REGION Network 357
   RUNG wire#powerrail
      Contact( "DuplicateCarrierfound" )
      Coil( "Carrier_17_Duplicate_Carrier_Fault" )
   END_RUNG
   // the same network as SCL:
   "Carrier_17_Duplicate_Carrier_Fault" := "DuplicateCarrierfound";
END_REGION

REGION Network 358
   RUNG wire#powerrail
      Contact( "EMS".Carrier[17].SDC_OUT.Faults.MotionOnFault )
      Coil( "Carrier_17_Motion_On_Fault" )
   END_RUNG
   // the same network as SCL:
   "Carrier_17_Motion_On_Fault" := "EMS".Carrier[17].SDC_OUT.Faults.MotionOnFault;
END_REGION

REGION Network 359
   RUNG wire#powerrail
      Contact( "EMS".Carrier[17].SDC_OUT.Faults.MotionOffFault )
      Coil( "Carrier_17_Motion_Off_Fault" )
   END_RUNG
   // the same network as SCL:
   "Carrier_17_Motion_Off_Fault" := "EMS".Carrier[17].SDC_OUT.Faults.MotionOffFault;
END_REGION

REGION Network 360
   RUNG wire#powerrail
      Contact( "EMS".Carrier[17].SDC_OUT.Faults.CarrierSpacingFault )
      Coil( "Carrier_17_Carrier_Spacing_Fault" )
   END_RUNG
   // the same network as SCL:
   "Carrier_17_Carrier_Spacing_Fault" := "EMS".Carrier[17].SDC_OUT.Faults.CarrierSpacingFault;
END_REGION

REGION Network 361
   RUNG wire#powerrail
      Move(in := "EMS".Carrier[18].SDC_OUT.Zone, out1 => "Carrier_18_Carrier_In_Zone")
   END_RUNG
   // the same network as SCL:
   "Carrier_18_Carrier_In_Zone" := "EMS".Carrier[18].SDC_OUT.Zone;
END_REGION

REGION Network 362
   RUNG wire#powerrail
      Move(in := "EMS".Carrier[18].SDC_OUT.CarrierNum, out1 => "Carrier_18_Carrier_Number_Echo")
   END_RUNG
   // the same network as SCL:
   "Carrier_18_Carrier_Number_Echo" := "EMS".Carrier[18].SDC_OUT.CarrierNum;
END_REGION

REGION Network 363
   RUNG wire#powerrail
      Move(in := "EMS".Carrier[18].SDC_OUT.CarrierPosition, out1 => "Carrier_18_Carrier_Position_Echo")
   END_RUNG
   // the same network as SCL:
   "Carrier_18_Carrier_Position_Echo" := "EMS".Carrier[18].SDC_OUT.CarrierPosition;
END_REGION

REGION Network 364
   RUNG wire#powerrail
      Move(in := "EMS".Carrier[18].SDC_OUT.NextCarrierNum, out1 => "Carrier_18_Next_Carrier_Number")
   END_RUNG
   // the same network as SCL:
   "Carrier_18_Next_Carrier_Number" := "EMS".Carrier[18].SDC_OUT.NextCarrierNum;
END_REGION

REGION Network 365
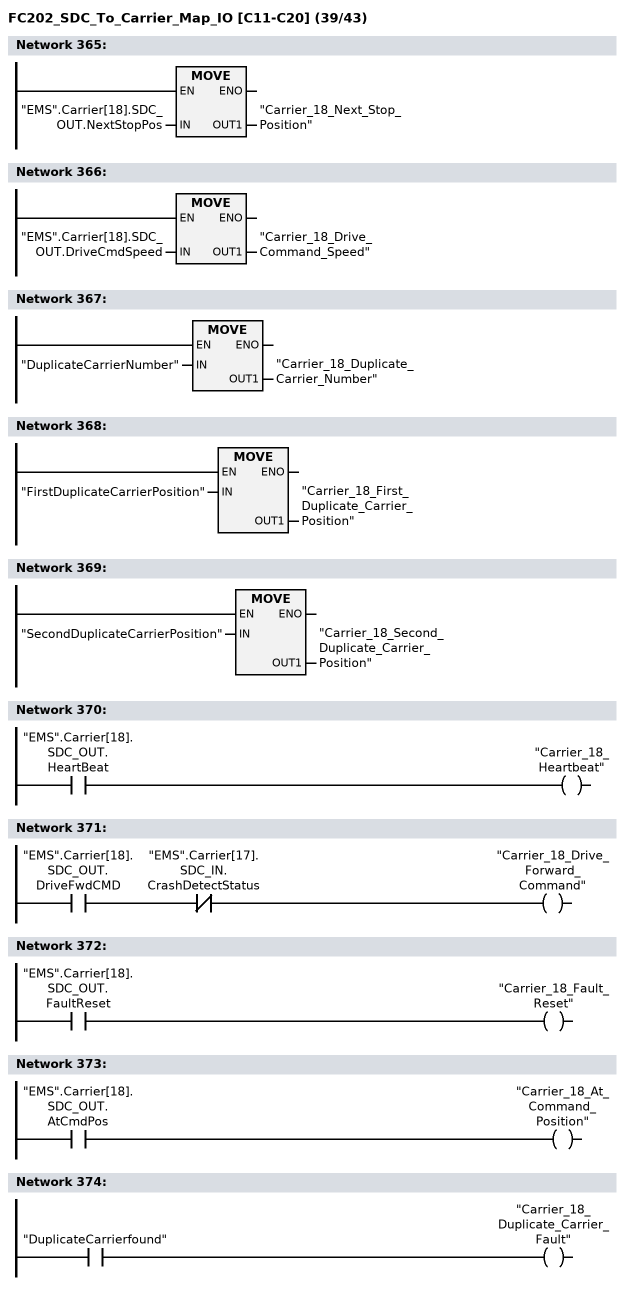
   RUNG wire#powerrail
      Move(in := "EMS".Carrier[18].SDC_OUT.NextStopPos, out1 => "Carrier_18_Next_Stop_Position")
   END_RUNG
   // the same network as SCL:
   "Carrier_18_Next_Stop_Position" := "EMS".Carrier[18].SDC_OUT.NextStopPos;
END_REGION

REGION Network 366
   RUNG wire#powerrail
      Move(in := "EMS".Carrier[18].SDC_OUT.DriveCmdSpeed, out1 => "Carrier_18_Drive_Command_Speed")
   END_RUNG
   // the same network as SCL:
   "Carrier_18_Drive_Command_Speed" := "EMS".Carrier[18].SDC_OUT.DriveCmdSpeed;
END_REGION

REGION Network 367
   RUNG wire#powerrail
      Move(in := "DuplicateCarrierNumber", out1 => "Carrier_18_Duplicate_Carrier_Number")
   END_RUNG
   // the same network as SCL:
   "Carrier_18_Duplicate_Carrier_Number" := "DuplicateCarrierNumber";
END_REGION

REGION Network 368
   RUNG wire#powerrail
      Move(in := "FirstDuplicateCarrierPosition", out1 => "Carrier_18_First_Duplicate_Carrier_Position")
   END_RUNG
   // the same network as SCL:
   "Carrier_18_First_Duplicate_Carrier_Position" := "FirstDuplicateCarrierPosition";
END_REGION

REGION Network 369
   RUNG wire#powerrail
      Move(in := "SecondDuplicateCarrierPosition", out1 => "Carrier_18_Second_Duplicate_Carrier_Position")
   END_RUNG
   // the same network as SCL:
   "Carrier_18_Second_Duplicate_Carrier_Position" := "SecondDuplicateCarrierPosition";
END_REGION

REGION Network 370
   RUNG wire#powerrail
      Contact( "EMS".Carrier[18].SDC_OUT.HeartBeat )
      Coil( "Carrier_18_Heartbeat" )
   END_RUNG
   // the same network as SCL:
   "Carrier_18_Heartbeat" := "EMS".Carrier[18].SDC_OUT.HeartBeat;
END_REGION

REGION Network 371
   RUNG wire#powerrail
      Contact( "EMS".Carrier[18].SDC_OUT.DriveFwdCMD )
      I_Contact( "EMS".Carrier[17].SDC_IN.CrashDetectStatus )
      Coil( "Carrier_18_Drive_Forward_Command" )
   END_RUNG
   // the same network as SCL:
   "Carrier_18_Drive_Forward_Command" := "EMS".Carrier[18].SDC_OUT.DriveFwdCMD AND NOT "EMS".Carrier[17].SDC_IN.CrashDetectStatus;
END_REGION

REGION Network 372
   RUNG wire#powerrail
      Contact( "EMS".Carrier[18].SDC_OUT.FaultReset )
      Coil( "Carrier_18_Fault_Reset" )
   END_RUNG
   // the same network as SCL:
   "Carrier_18_Fault_Reset" := "EMS".Carrier[18].SDC_OUT.FaultReset;
END_REGION

REGION Network 373
   RUNG wire#powerrail
      Contact( "EMS".Carrier[18].SDC_OUT.AtCmdPos )
      Coil( "Carrier_18_At_Command_Position" )
   END_RUNG
   // the same network as SCL:
   "Carrier_18_At_Command_Position" := "EMS".Carrier[18].SDC_OUT.AtCmdPos;
END_REGION

REGION Network 374
   RUNG wire#powerrail
      Contact( "DuplicateCarrierfound" )
      Coil( "Carrier_18_Duplicate_Carrier_Fault" )
   END_RUNG
   // the same network as SCL:
   "Carrier_18_Duplicate_Carrier_Fault" := "DuplicateCarrierfound";
END_REGION

REGION Network 375
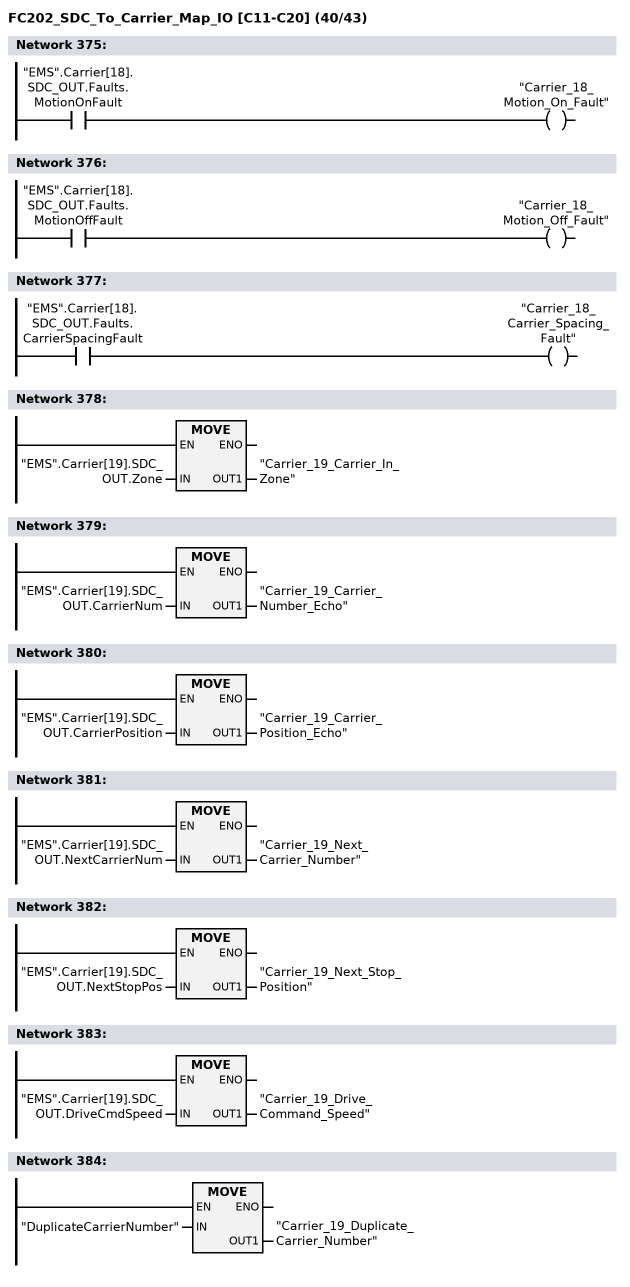
   RUNG wire#powerrail
      Contact( "EMS".Carrier[18].SDC_OUT.Faults.MotionOnFault )
      Coil( "Carrier_18_Motion_On_Fault" )
   END_RUNG
   // the same network as SCL:
   "Carrier_18_Motion_On_Fault" := "EMS".Carrier[18].SDC_OUT.Faults.MotionOnFault;
END_REGION

REGION Network 376
   RUNG wire#powerrail
      Contact( "EMS".Carrier[18].SDC_OUT.Faults.MotionOffFault )
      Coil( "Carrier_18_Motion_Off_Fault" )
   END_RUNG
   // the same network as SCL:
   "Carrier_18_Motion_Off_Fault" := "EMS".Carrier[18].SDC_OUT.Faults.MotionOffFault;
END_REGION

REGION Network 377
   RUNG wire#powerrail
      Contact( "EMS".Carrier[18].SDC_OUT.Faults.CarrierSpacingFault )
      Coil( "Carrier_18_Carrier_Spacing_Fault" )
   END_RUNG
   // the same network as SCL:
   "Carrier_18_Carrier_Spacing_Fault" := "EMS".Carrier[18].SDC_OUT.Faults.CarrierSpacingFault;
END_REGION

REGION Network 378
   RUNG wire#powerrail
      Move(in := "EMS".Carrier[19].SDC_OUT.Zone, out1 => "Carrier_19_Carrier_In_Zone")
   END_RUNG
   // the same network as SCL:
   "Carrier_19_Carrier_In_Zone" := "EMS".Carrier[19].SDC_OUT.Zone;
END_REGION

REGION Network 379
   RUNG wire#powerrail
      Move(in := "EMS".Carrier[19].SDC_OUT.CarrierNum, out1 => "Carrier_19_Carrier_Number_Echo")
   END_RUNG
   // the same network as SCL:
   "Carrier_19_Carrier_Number_Echo" := "EMS".Carrier[19].SDC_OUT.CarrierNum;
END_REGION

REGION Network 380
   RUNG wire#powerrail
      Move(in := "EMS".Carrier[19].SDC_OUT.CarrierPosition, out1 => "Carrier_19_Carrier_Position_Echo")
   END_RUNG
   // the same network as SCL:
   "Carrier_19_Carrier_Position_Echo" := "EMS".Carrier[19].SDC_OUT.CarrierPosition;
END_REGION

REGION Network 381
   RUNG wire#powerrail
      Move(in := "EMS".Carrier[19].SDC_OUT.NextCarrierNum, out1 => "Carrier_19_Next_Carrier_Number")
   END_RUNG
   // the same network as SCL:
   "Carrier_19_Next_Carrier_Number" := "EMS".Carrier[19].SDC_OUT.NextCarrierNum;
END_REGION

REGION Network 382
   RUNG wire#powerrail
      Move(in := "EMS".Carrier[19].SDC_OUT.NextStopPos, out1 => "Carrier_19_Next_Stop_Position")
   END_RUNG
   // the same network as SCL:
   "Carrier_19_Next_Stop_Position" := "EMS".Carrier[19].SDC_OUT.NextStopPos;
END_REGION

REGION Network 383
   RUNG wire#powerrail
      Move(in := "EMS".Carrier[19].SDC_OUT.DriveCmdSpeed, out1 => "Carrier_19_Drive_Command_Speed")
   END_RUNG
   // the same network as SCL:
   "Carrier_19_Drive_Command_Speed" := "EMS".Carrier[19].SDC_OUT.DriveCmdSpeed;
END_REGION

REGION Network 384
   RUNG wire#powerrail
      Move(in := "DuplicateCarrierNumber", out1 => "Carrier_19_Duplicate_Carrier_Number")
   END_RUNG
   // the same network as SCL:
   "Carrier_19_Duplicate_Carrier_Number" := "DuplicateCarrierNumber";
END_REGION

REGION Network 385
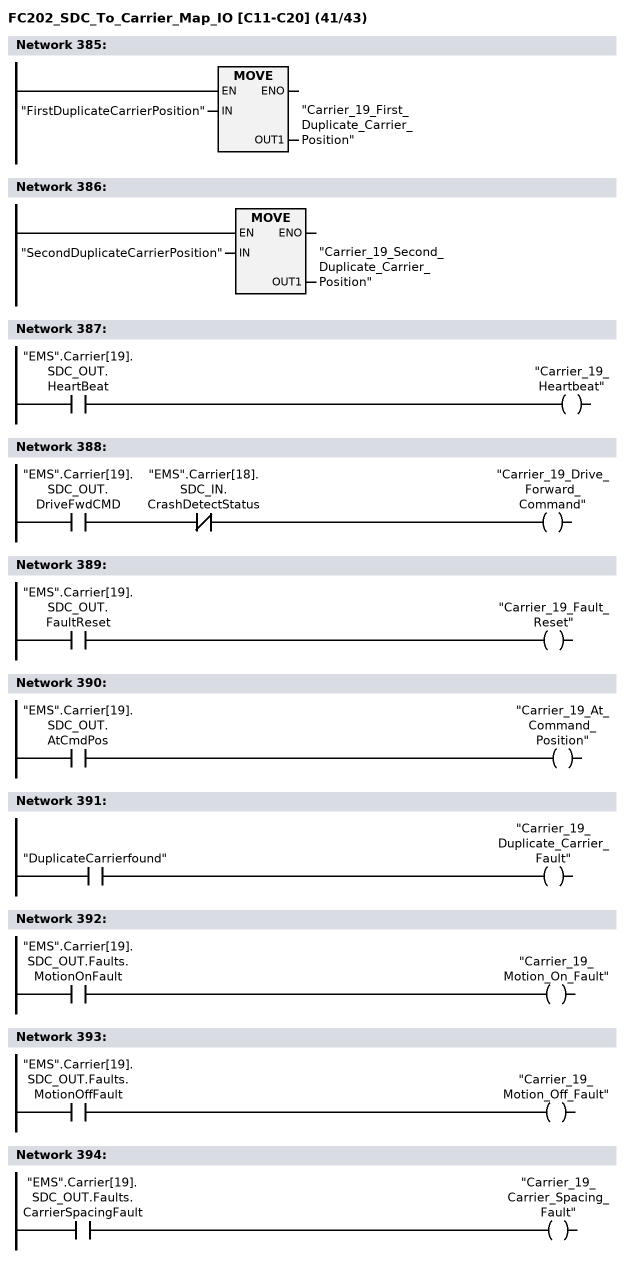
   RUNG wire#powerrail
      Move(in := "FirstDuplicateCarrierPosition", out1 => "Carrier_19_First_Duplicate_Carrier_Position")
   END_RUNG
   // the same network as SCL:
   "Carrier_19_First_Duplicate_Carrier_Position" := "FirstDuplicateCarrierPosition";
END_REGION

REGION Network 386
   RUNG wire#powerrail
      Move(in := "SecondDuplicateCarrierPosition", out1 => "Carrier_19_Second_Duplicate_Carrier_Position")
   END_RUNG
   // the same network as SCL:
   "Carrier_19_Second_Duplicate_Carrier_Position" := "SecondDuplicateCarrierPosition";
END_REGION

REGION Network 387
   RUNG wire#powerrail
      Contact( "EMS".Carrier[19].SDC_OUT.HeartBeat )
      Coil( "Carrier_19_Heartbeat" )
   END_RUNG
   // the same network as SCL:
   "Carrier_19_Heartbeat" := "EMS".Carrier[19].SDC_OUT.HeartBeat;
END_REGION

REGION Network 388
   RUNG wire#powerrail
      Contact( "EMS".Carrier[19].SDC_OUT.DriveFwdCMD )
      I_Contact( "EMS".Carrier[18].SDC_IN.CrashDetectStatus )
      Coil( "Carrier_19_Drive_Forward_Command" )
   END_RUNG
   // the same network as SCL:
   "Carrier_19_Drive_Forward_Command" := "EMS".Carrier[19].SDC_OUT.DriveFwdCMD AND NOT "EMS".Carrier[18].SDC_IN.CrashDetectStatus;
END_REGION

REGION Network 389
   RUNG wire#powerrail
      Contact( "EMS".Carrier[19].SDC_OUT.FaultReset )
      Coil( "Carrier_19_Fault_Reset" )
   END_RUNG
   // the same network as SCL:
   "Carrier_19_Fault_Reset" := "EMS".Carrier[19].SDC_OUT.FaultReset;
END_REGION

REGION Network 390
   RUNG wire#powerrail
      Contact( "EMS".Carrier[19].SDC_OUT.AtCmdPos )
      Coil( "Carrier_19_At_Command_Position" )
   END_RUNG
   // the same network as SCL:
   "Carrier_19_At_Command_Position" := "EMS".Carrier[19].SDC_OUT.AtCmdPos;
END_REGION

REGION Network 391
   RUNG wire#powerrail
      Contact( "DuplicateCarrierfound" )
      Coil( "Carrier_19_Duplicate_Carrier_Fault" )
   END_RUNG
   // the same network as SCL:
   "Carrier_19_Duplicate_Carrier_Fault" := "DuplicateCarrierfound";
END_REGION

REGION Network 392
   RUNG wire#powerrail
      Contact( "EMS".Carrier[19].SDC_OUT.Faults.MotionOnFault )
      Coil( "Carrier_19_Motion_On_Fault" )
   END_RUNG
   // the same network as SCL:
   "Carrier_19_Motion_On_Fault" := "EMS".Carrier[19].SDC_OUT.Faults.MotionOnFault;
END_REGION

REGION Network 393
   RUNG wire#powerrail
      Contact( "EMS".Carrier[19].SDC_OUT.Faults.MotionOffFault )
      Coil( "Carrier_19_Motion_Off_Fault" )
   END_RUNG
   // the same network as SCL:
   "Carrier_19_Motion_Off_Fault" := "EMS".Carrier[19].SDC_OUT.Faults.MotionOffFault;
END_REGION

REGION Network 394
   RUNG wire#powerrail
      Contact( "EMS".Carrier[19].SDC_OUT.Faults.CarrierSpacingFault )
      Coil( "Carrier_19_Carrier_Spacing_Fault" )
   END_RUNG
   // the same network as SCL:
   "Carrier_19_Carrier_Spacing_Fault" := "EMS".Carrier[19].SDC_OUT.Faults.CarrierSpacingFault;
END_REGION

REGION Network 395
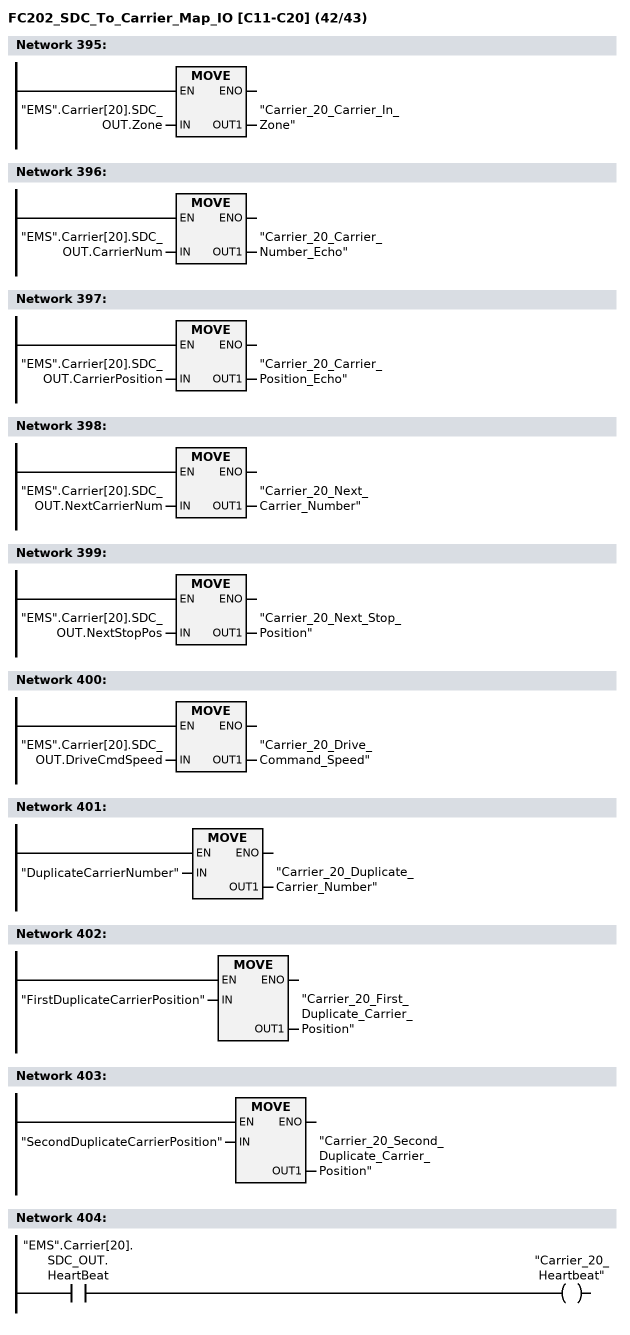
   RUNG wire#powerrail
      Move(in := "EMS".Carrier[20].SDC_OUT.Zone, out1 => "Carrier_20_Carrier_In_Zone")
   END_RUNG
   // the same network as SCL:
   "Carrier_20_Carrier_In_Zone" := "EMS".Carrier[20].SDC_OUT.Zone;
END_REGION

REGION Network 396
   RUNG wire#powerrail
      Move(in := "EMS".Carrier[20].SDC_OUT.CarrierNum, out1 => "Carrier_20_Carrier_Number_Echo")
   END_RUNG
   // the same network as SCL:
   "Carrier_20_Carrier_Number_Echo" := "EMS".Carrier[20].SDC_OUT.CarrierNum;
END_REGION

REGION Network 397
   RUNG wire#powerrail
      Move(in := "EMS".Carrier[20].SDC_OUT.CarrierPosition, out1 => "Carrier_20_Carrier_Position_Echo")
   END_RUNG
   // the same network as SCL:
   "Carrier_20_Carrier_Position_Echo" := "EMS".Carrier[20].SDC_OUT.CarrierPosition;
END_REGION

REGION Network 398
   RUNG wire#powerrail
      Move(in := "EMS".Carrier[20].SDC_OUT.NextCarrierNum, out1 => "Carrier_20_Next_Carrier_Number")
   END_RUNG
   // the same network as SCL:
   "Carrier_20_Next_Carrier_Number" := "EMS".Carrier[20].SDC_OUT.NextCarrierNum;
END_REGION

REGION Network 399
   RUNG wire#powerrail
      Move(in := "EMS".Carrier[20].SDC_OUT.NextStopPos, out1 => "Carrier_20_Next_Stop_Position")
   END_RUNG
   // the same network as SCL:
   "Carrier_20_Next_Stop_Position" := "EMS".Carrier[20].SDC_OUT.NextStopPos;
END_REGION

REGION Network 400
   RUNG wire#powerrail
      Move(in := "EMS".Carrier[20].SDC_OUT.DriveCmdSpeed, out1 => "Carrier_20_Drive_Command_Speed")
   END_RUNG
   // the same network as SCL:
   "Carrier_20_Drive_Command_Speed" := "EMS".Carrier[20].SDC_OUT.DriveCmdSpeed;
END_REGION

REGION Network 401
   RUNG wire#powerrail
      Move(in := "DuplicateCarrierNumber", out1 => "Carrier_20_Duplicate_Carrier_Number")
   END_RUNG
   // the same network as SCL:
   "Carrier_20_Duplicate_Carrier_Number" := "DuplicateCarrierNumber";
END_REGION

REGION Network 402
   RUNG wire#powerrail
      Move(in := "FirstDuplicateCarrierPosition", out1 => "Carrier_20_First_Duplicate_Carrier_Position")
   END_RUNG
   // the same network as SCL:
   "Carrier_20_First_Duplicate_Carrier_Position" := "FirstDuplicateCarrierPosition";
END_REGION

REGION Network 403
   RUNG wire#powerrail
      Move(in := "SecondDuplicateCarrierPosition", out1 => "Carrier_20_Second_Duplicate_Carrier_Position")
   END_RUNG
   // the same network as SCL:
   "Carrier_20_Second_Duplicate_Carrier_Position" := "SecondDuplicateCarrierPosition";
END_REGION

REGION Network 404
   RUNG wire#powerrail
      Contact( "EMS".Carrier[20].SDC_OUT.HeartBeat )
      Coil( "Carrier_20_Heartbeat" )
   END_RUNG
   // the same network as SCL:
   "Carrier_20_Heartbeat" := "EMS".Carrier[20].SDC_OUT.HeartBeat;
END_REGION

REGION Network 405
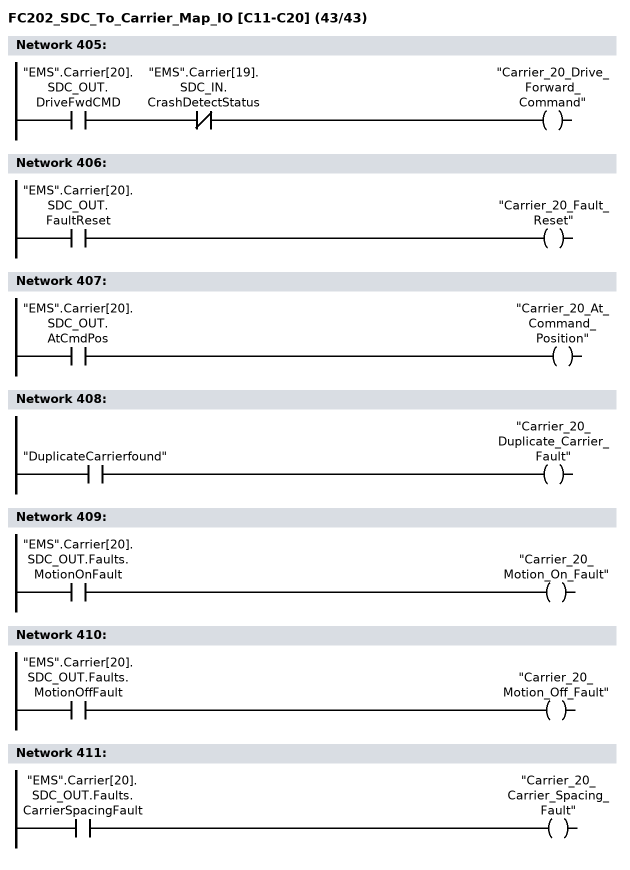
   RUNG wire#powerrail
      Contact( "EMS".Carrier[20].SDC_OUT.DriveFwdCMD )
      I_Contact( "EMS".Carrier[19].SDC_IN.CrashDetectStatus )
      Coil( "Carrier_20_Drive_Forward_Command" )
   END_RUNG
   // the same network as SCL:
   "Carrier_20_Drive_Forward_Command" := "EMS".Carrier[20].SDC_OUT.DriveFwdCMD AND NOT "EMS".Carrier[19].SDC_IN.CrashDetectStatus;
END_REGION

REGION Network 406
   RUNG wire#powerrail
      Contact( "EMS".Carrier[20].SDC_OUT.FaultReset )
      Coil( "Carrier_20_Fault_Reset" )
   END_RUNG
   // the same network as SCL:
   "Carrier_20_Fault_Reset" := "EMS".Carrier[20].SDC_OUT.FaultReset;
END_REGION

REGION Network 407
   RUNG wire#powerrail
      Contact( "EMS".Carrier[20].SDC_OUT.AtCmdPos )
      Coil( "Carrier_20_At_Command_Position" )
   END_RUNG
   // the same network as SCL:
   "Carrier_20_At_Command_Position" := "EMS".Carrier[20].SDC_OUT.AtCmdPos;
END_REGION

REGION Network 408
   RUNG wire#powerrail
      Contact( "DuplicateCarrierfound" )
      Coil( "Carrier_20_Duplicate_Carrier_Fault" )
   END_RUNG
   // the same network as SCL:
   "Carrier_20_Duplicate_Carrier_Fault" := "DuplicateCarrierfound";
END_REGION

REGION Network 409
   RUNG wire#powerrail
      Contact( "EMS".Carrier[20].SDC_OUT.Faults.MotionOnFault )
      Coil( "Carrier_20_Motion_On_Fault" )
   END_RUNG
   // the same network as SCL:
   "Carrier_20_Motion_On_Fault" := "EMS".Carrier[20].SDC_OUT.Faults.MotionOnFault;
END_REGION

REGION Network 410
   RUNG wire#powerrail
      Contact( "EMS".Carrier[20].SDC_OUT.Faults.MotionOffFault )
      Coil( "Carrier_20_Motion_Off_Fault" )
   END_RUNG
   // the same network as SCL:
   "Carrier_20_Motion_Off_Fault" := "EMS".Carrier[20].SDC_OUT.Faults.MotionOffFault;
END_REGION

REGION Network 411
   RUNG wire#powerrail
      Contact( "EMS".Carrier[20].SDC_OUT.Faults.CarrierSpacingFault )
      Coil( "Carrier_20_Carrier_Spacing_Fault" )
   END_RUNG
   // the same network as SCL:
   "Carrier_20_Carrier_Spacing_Fault" := "EMS".Carrier[20].SDC_OUT.Faults.CarrierSpacingFault;
END_REGION
END_FUNCTION

FUNCTION "FC203_SDC_To_Carrier_Map_IO [C21-C30]" : Void   // FC203, LAD
{ S7_Optimized_Access := 'TRUE' }
VERSION : 0.1
BEGIN

REGION Network 1
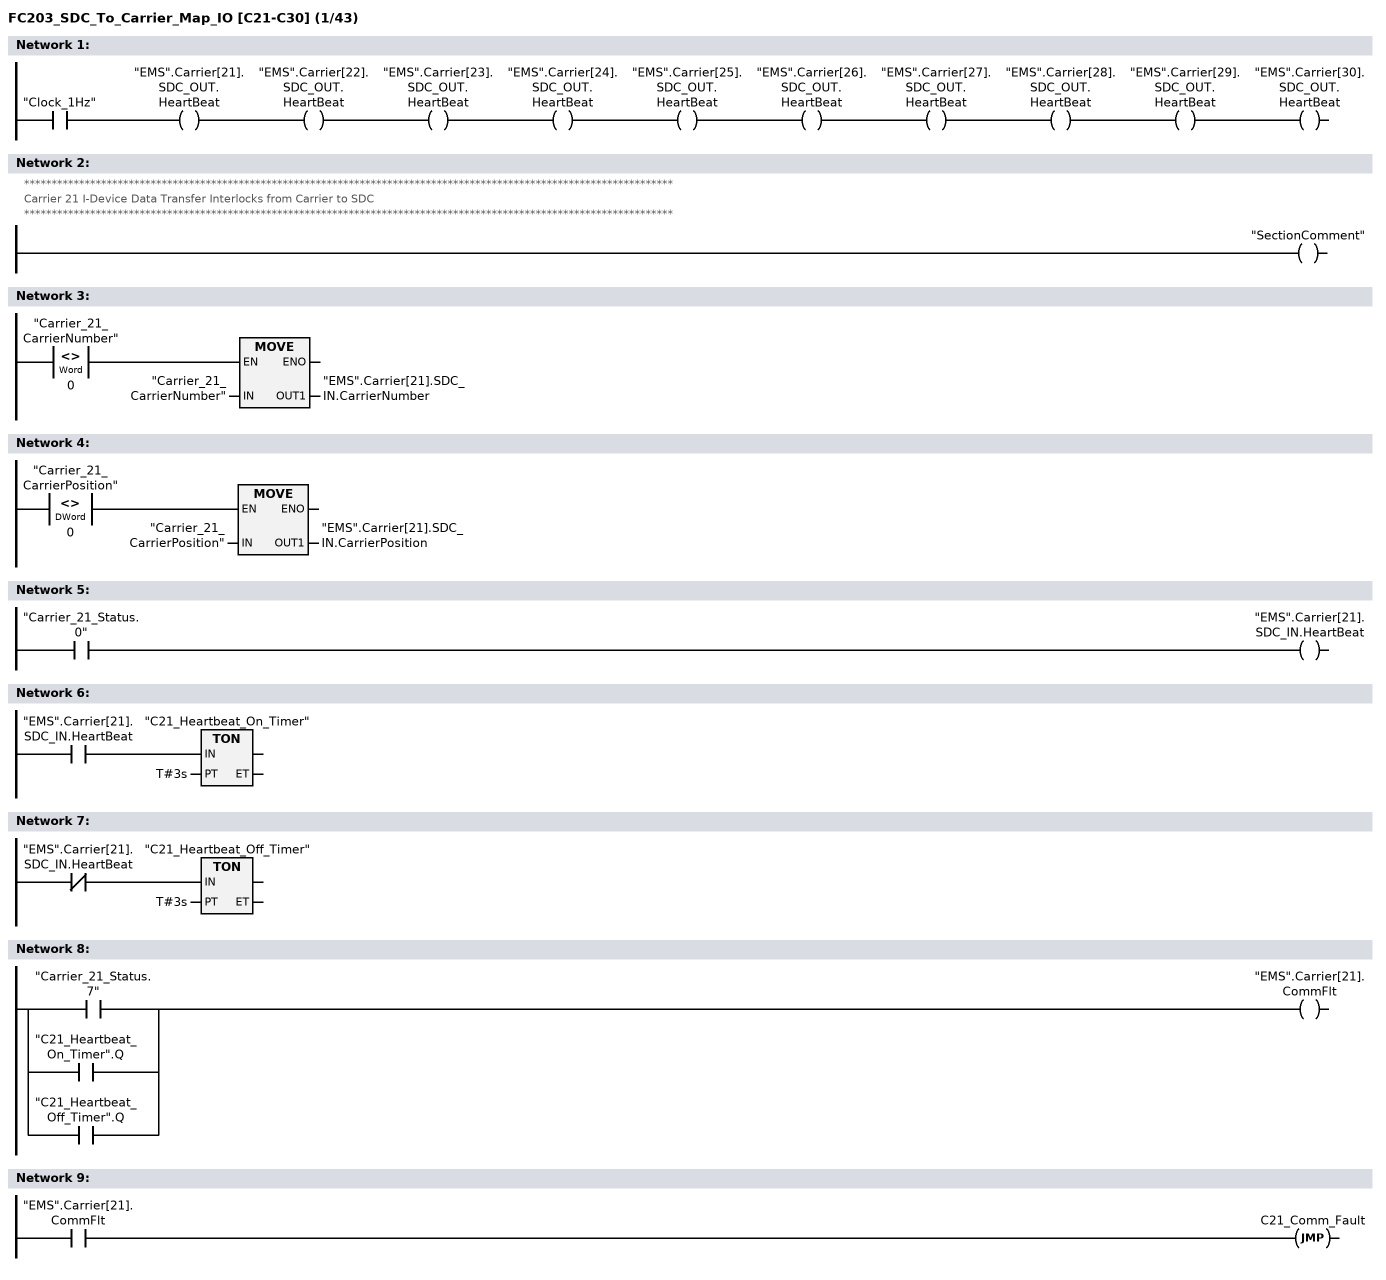
   RUNG wire#powerrail
      Contact( "Clock_1Hz" )
      Coil( "EMS".Carrier[21].SDC_OUT.HeartBeat )
      Coil( "EMS".Carrier[22].SDC_OUT.HeartBeat )
      Coil( "EMS".Carrier[23].SDC_OUT.HeartBeat )
      Coil( "EMS".Carrier[24].SDC_OUT.HeartBeat )
      Coil( "EMS".Carrier[25].SDC_OUT.HeartBeat )
      Coil( "EMS".Carrier[26].SDC_OUT.HeartBeat )
      Coil( "EMS".Carrier[27].SDC_OUT.HeartBeat )
      Coil( "EMS".Carrier[28].SDC_OUT.HeartBeat )
      Coil( "EMS".Carrier[29].SDC_OUT.HeartBeat )
      Coil( "EMS".Carrier[30].SDC_OUT.HeartBeat )
   END_RUNG
   // the same network as SCL:
   "EMS".Carrier[21].SDC_OUT.HeartBeat := "Clock_1Hz";
   "EMS".Carrier[22].SDC_OUT.HeartBeat := "Clock_1Hz";
   "EMS".Carrier[23].SDC_OUT.HeartBeat := "Clock_1Hz";
   "EMS".Carrier[24].SDC_OUT.HeartBeat := "Clock_1Hz";
   "EMS".Carrier[25].SDC_OUT.HeartBeat := "Clock_1Hz";
   "EMS".Carrier[26].SDC_OUT.HeartBeat := "Clock_1Hz";
   "EMS".Carrier[27].SDC_OUT.HeartBeat := "Clock_1Hz";
   "EMS".Carrier[28].SDC_OUT.HeartBeat := "Clock_1Hz";
   "EMS".Carrier[29].SDC_OUT.HeartBeat := "Clock_1Hz";
   "EMS".Carrier[30].SDC_OUT.HeartBeat := "Clock_1Hz";
END_REGION

REGION Network 2
   // **********************************************************************************************************************
   // 
   // Carrier 21 I-Device Data Transfer Interlocks from Carrier to SDC
   // 
   // **********************************************************************************************************************
   RUNG wire#powerrail
      Coil( "SectionComment" )
   END_RUNG
   // the same network as SCL:
   "SectionComment" := TRUE;
END_REGION

REGION Network 3
   RUNG wire#powerrail
      { S7_Templates := "SrcType := Word" } NE_Contact(in1 := "Carrier_21_CarrierNumber", in2 := 0)
      Move(in := "Carrier_21_CarrierNumber", out1 => "EMS".Carrier[21].SDC_IN.CarrierNumber)
   END_RUNG
   // the same network as SCL:
   IF "Carrier_21_CarrierNumber" <> 0 THEN
       "EMS".Carrier[21].SDC_IN.CarrierNumber := "Carrier_21_CarrierNumber";
   END_IF;
END_REGION

REGION Network 4
   RUNG wire#powerrail
      { S7_Templates := "SrcType := DWord" } NE_Contact(in1 := "Carrier_21_CarrierPosition", in2 := 0)
      Move(in := "Carrier_21_CarrierPosition", out1 => "EMS".Carrier[21].SDC_IN.CarrierPosition)
   END_RUNG
   // the same network as SCL:
   IF "Carrier_21_CarrierPosition" <> 0 THEN
       "EMS".Carrier[21].SDC_IN.CarrierPosition := "Carrier_21_CarrierPosition";
   END_IF;
END_REGION

REGION Network 5
   RUNG wire#powerrail
      Contact( "Carrier_21_Status.0" )
      Coil( "EMS".Carrier[21].SDC_IN.HeartBeat )
   END_RUNG
   // the same network as SCL:
   "EMS".Carrier[21].SDC_IN.HeartBeat := "Carrier_21_Status.0";
END_REGION

REGION Network 6
   "C21_Heartbeat_On_Timer".TON(IN := "EMS".Carrier[21].SDC_IN.HeartBeat, PT := T#3s);
END_REGION

REGION Network 7
   "C21_Heartbeat_Off_Timer".TON(IN := NOT "EMS".Carrier[21].SDC_IN.HeartBeat, PT := T#3s);
END_REGION

REGION Network 8
   RUNG wire#powerrail
      Contact( "Carrier_21_Status.7" )
      wire#w1
      Coil( "EMS".Carrier[21].CommFlt )
   END_RUNG
   RUNG wire#powerrail
      Contact( "C21_Heartbeat_On_Timer".Q )
   END_RUNG wire#w1
   RUNG wire#powerrail
      Contact( "C21_Heartbeat_Off_Timer".Q )
   END_RUNG wire#w1
   // the same network as SCL:
   "EMS".Carrier[21].CommFlt := "Carrier_21_Status.7" OR "C21_Heartbeat_On_Timer".Q OR "C21_Heartbeat_Off_Timer".Q;
END_REGION

REGION Network 9
   RUNG wire#powerrail
      Contact( "EMS".Carrier[21].CommFlt )
      JumpCoil( C21_Comm_Fault )
   END_RUNG
   // the same network as SCL:
   IF "EMS".Carrier[21].CommFlt THEN GOTO C21_Comm_Fault; END_IF;
END_REGION

REGION Network 10
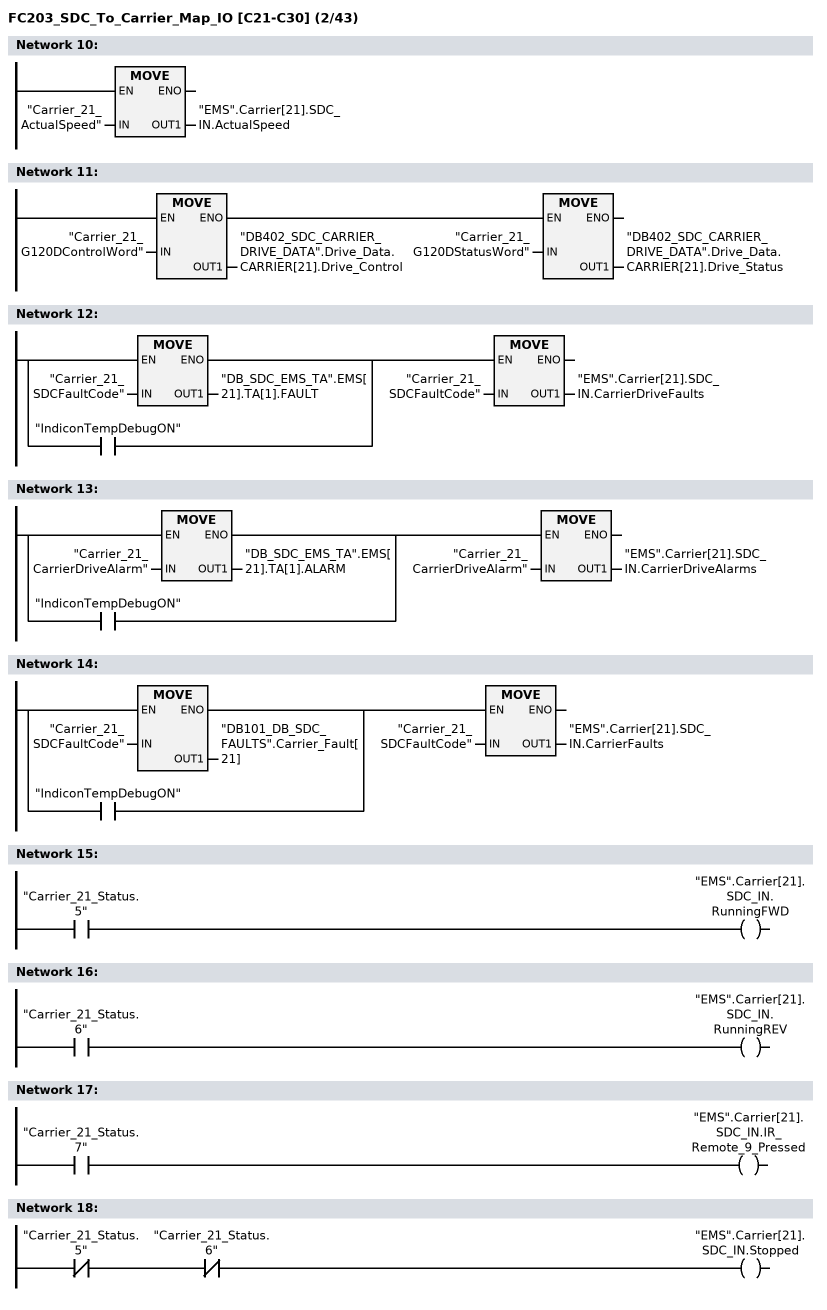
   RUNG wire#powerrail
      Move(in := "Carrier_21_ActualSpeed", out1 => "EMS".Carrier[21].SDC_IN.ActualSpeed)
   END_RUNG
   // the same network as SCL:
   "EMS".Carrier[21].SDC_IN.ActualSpeed := "Carrier_21_ActualSpeed";
END_REGION

REGION Network 11
   RUNG wire#powerrail
      Move(in := "Carrier_21_G120DControlWord", out1 => "DB402_SDC_CARRIER_DRIVE_DATA".Drive_Data.CARRIER[21].Drive_Control)
      Move(in := "Carrier_21_G120DStatusWord", out1 => "DB402_SDC_CARRIER_DRIVE_DATA".Drive_Data.CARRIER[21].Drive_Status)
   END_RUNG
   // the same network as SCL:
   "DB402_SDC_CARRIER_DRIVE_DATA".Drive_Data.CARRIER[21].Drive_Control := "Carrier_21_G120DControlWord";
   "DB402_SDC_CARRIER_DRIVE_DATA".Drive_Data.CARRIER[21].Drive_Status := "Carrier_21_G120DStatusWord";
END_REGION

REGION Network 12
   RUNG wire#powerrail
      Move(in := "Carrier_21_SDCFaultCode", out1 => "DB_SDC_EMS_TA".EMS[21].TA[1].FAULT)
      wire#w1
      Move(in := "Carrier_21_SDCFaultCode", out1 => "EMS".Carrier[21].SDC_IN.CarrierDriveFaults)
   END_RUNG
   RUNG wire#powerrail
      Contact( "IndiconTempDebugON" )
   END_RUNG wire#w1
   // the same network as SCL:
   "DB_SDC_EMS_TA".EMS[21].TA[1].FAULT := "Carrier_21_SDCFaultCode";
   IF TRUE OR "IndiconTempDebugON" THEN
       "EMS".Carrier[21].SDC_IN.CarrierDriveFaults := "Carrier_21_SDCFaultCode";
   END_IF;
END_REGION

REGION Network 13
   RUNG wire#powerrail
      Move(in := "Carrier_21_CarrierDriveAlarm", out1 => "DB_SDC_EMS_TA".EMS[21].TA[1].ALARM)
      wire#w1
      Move(in := "Carrier_21_CarrierDriveAlarm", out1 => "EMS".Carrier[21].SDC_IN.CarrierDriveAlarms)
   END_RUNG
   RUNG wire#powerrail
      Contact( "IndiconTempDebugON" )
   END_RUNG wire#w1
   // the same network as SCL:
   "DB_SDC_EMS_TA".EMS[21].TA[1].ALARM := "Carrier_21_CarrierDriveAlarm";
   IF TRUE OR "IndiconTempDebugON" THEN
       "EMS".Carrier[21].SDC_IN.CarrierDriveAlarms := "Carrier_21_CarrierDriveAlarm";
   END_IF;
END_REGION

REGION Network 14
   RUNG wire#powerrail
      Move(in := "Carrier_21_SDCFaultCode", out1 => "DB101_DB_SDC_FAULTS".Carrier_Fault[21])
      wire#w1
      Move(in := "Carrier_21_SDCFaultCode", out1 => "EMS".Carrier[21].SDC_IN.CarrierFaults)
   END_RUNG
   RUNG wire#powerrail
      Contact( "IndiconTempDebugON" )
   END_RUNG wire#w1
   // the same network as SCL:
   "DB101_DB_SDC_FAULTS".Carrier_Fault[21] := "Carrier_21_SDCFaultCode";
   IF TRUE OR "IndiconTempDebugON" THEN
       "EMS".Carrier[21].SDC_IN.CarrierFaults := "Carrier_21_SDCFaultCode";
   END_IF;
END_REGION

REGION Network 15
   RUNG wire#powerrail
      Contact( "Carrier_21_Status.5" )
      Coil( "EMS".Carrier[21].SDC_IN.RunningFWD )
   END_RUNG
   // the same network as SCL:
   "EMS".Carrier[21].SDC_IN.RunningFWD := "Carrier_21_Status.5";
END_REGION

REGION Network 16
   RUNG wire#powerrail
      Contact( "Carrier_21_Status.6" )
      Coil( "EMS".Carrier[21].SDC_IN.RunningREV )
   END_RUNG
   // the same network as SCL:
   "EMS".Carrier[21].SDC_IN.RunningREV := "Carrier_21_Status.6";
END_REGION

REGION Network 17
   RUNG wire#powerrail
      Contact( "Carrier_21_Status.7" )
      Coil( "EMS".Carrier[21].SDC_IN.IR_Remote_9_Pressed )
   END_RUNG
   // the same network as SCL:
   "EMS".Carrier[21].SDC_IN.IR_Remote_9_Pressed := "Carrier_21_Status.7";
END_REGION

REGION Network 18
   RUNG wire#powerrail
      I_Contact( "Carrier_21_Status.5" )
      I_Contact( "Carrier_21_Status.6" )
      Coil( "EMS".Carrier[21].SDC_IN.Stopped )
   END_RUNG
   // the same network as SCL:
   "EMS".Carrier[21].SDC_IN.Stopped := NOT "Carrier_21_Status.5" AND NOT "Carrier_21_Status.6";
END_REGION

REGION Network 19
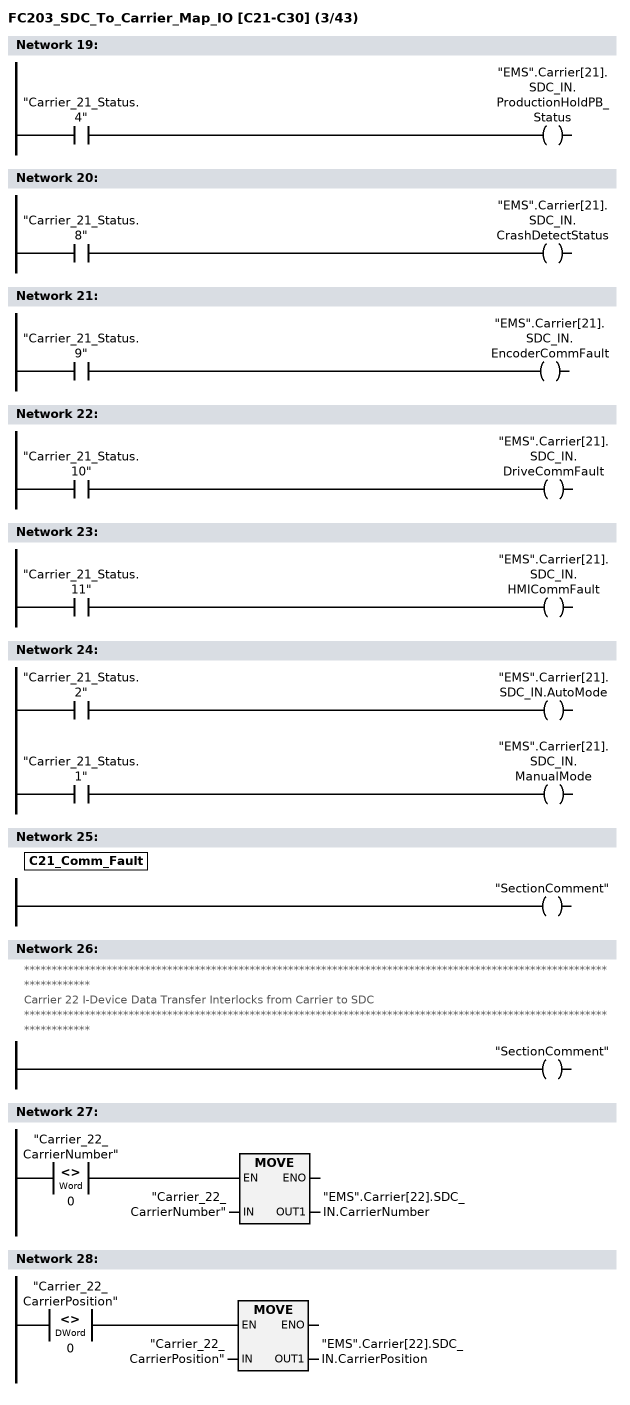
   RUNG wire#powerrail
      Contact( "Carrier_21_Status.4" )
      Coil( "EMS".Carrier[21].SDC_IN.ProductionHoldPB_Status )
   END_RUNG
   // the same network as SCL:
   "EMS".Carrier[21].SDC_IN.ProductionHoldPB_Status := "Carrier_21_Status.4";
END_REGION

REGION Network 20
   RUNG wire#powerrail
      Contact( "Carrier_21_Status.8" )
      Coil( "EMS".Carrier[21].SDC_IN.CrashDetectStatus )
   END_RUNG
   // the same network as SCL:
   "EMS".Carrier[21].SDC_IN.CrashDetectStatus := "Carrier_21_Status.8";
END_REGION
